// TIA Portal project "Linie_reciclare_paleti_mod" (V16)

(* hardware
DEVICE "S7-1200 station_1"  S7-1200 Station
   slot 0: "Rack_0"  S7-1200 Rack  Rack  V1.0
   slot 1: "150A19"  CPU 1214C DC/DC/Rly  6ES7 214-1HG40-0XB0  V4.4
   slot 2: "150A1101"  SM 1221 DI8 x 24VDC  6ES7 221-1BF30-0XB0  V1.0
   slot 3: "150A1102"  SM 1221 DI8 x 24VDC  6ES7 221-1BF30-0XB0  V1.0
   slot 4: "150A1103"  6ES7 221-1BH32-0XB0  V2.0
   slot 5: "150A1104"  6ES7 221-1BH32-0XB0  V2.0
   slot 6: "150A1105"  6ES7 221-1BH32-0XB0  V2.0
   slot 7: "150A1201"  SM 1222 DQ8 x relay  6ES7 222-1HF32-0XB0  V2.0
   slot 8: "150A1202"  SM 1222 DQ8 x relay  6ES7 222-1HF32-0XB0  V2.0
   slot 9: "150A1203"  SM 1222 DQ16 x relay  6ES7 222-1HH32-0XB0  V2.0
DEVICE "Master_Destacker"  GSD.Device.PN
   slot 0: "Rack"  Rack  V1.0
   slot 0: "Master_Destacker"  AL1100  AL1100
      slot 0: "AL1100"  AL1100
      slot 1: "X1"  X1
         slot 1: "Port 1"  Port 1
         slot 2: "Port 2"  Port 2
      slot 1: "4 Ports_1"  4 Ports  AL1100
         slot 0: "IO-Link Master"  IO-Link Master
   slot 1: "AL2401_IO-Link In  4 Byte + PQI"  IO-Link In  4 Byte + PQI
   slot 2: "AL2401_IO-Link In  4 Byte + PQI_1"  IO-Link In  4 Byte + PQI
   slot 3: "AL2330_IO-Link In/Out  8/ 8 Byte + PQI"  IO-Link In/Out  8/ 8 Byte + PQI
   slot 4: "IO-Link In/Out  2/ 2 Byte + PQI"  IO-Link In/Out  2/ 2 Byte + PQI
DEVICE "Master_Stacker"  GSD.Device.PN
   slot 0: "Rack"  Rack  V1.0
   slot 0: "Master_Stacker"  AL1100  AL1100
      slot 0: "AL1100"  AL1100
      slot 1: "X1"  X1
         slot 1: "Port 1"  Port 1
         slot 2: "Port 2"  Port 2
      slot 1: "4 Ports_1"  4 Ports  AL1100
         slot 0: "IO-Link Master"  IO-Link Master
   slot 1: "IO-Link In  4 Byte + PQI"  IO-Link In  4 Byte + PQI
   slot 2: "IO-Link In  4 Byte + PQI_1"  IO-Link In  4 Byte + PQI
   slot 3: "IO-Link In/Out  8/ 8 Byte + PQI"  IO-Link In/Out  8/ 8 Byte + PQI
   slot 4: "IO-Link In/Out  2/ 2 Byte + PQI"  IO-Link In/Out  2/ 2 Byte + PQI
DEVICE "HMI_1"  KTP700 Basic PN
   slot 0: "HMI_1"  KTP700 Basic PN  6AV2 123-2GB03-0AX0  16.0.0.0
   slot 1: "HMI_RT_1"  KTP700 Basic PN  6AV2 123-2GB03-0AX0  16.0.0.0
   slot 5: "HMI_1.IE_CP_1"  PROFINET Interface  16.0.0.0
      slot 1: "PROFINET Interface_1"  PROFINET Interface
         slot 1: "Port_1"  Port
DEVICE "HMI_2"  KTP700 Basic PN
   slot 0: "HMI_1"  KTP700 Basic PN  6AV2 123-2GB03-0AX0  16.0.0.0
   slot 1: "HMI_RT_2"  KTP700 Basic PN  6AV2 123-2GB03-0AX0  16.0.0.0
   slot 5: "HMI_1.IE_CP_1"  PROFINET Interface  16.0.0.0
      slot 1: "PROFINET Interface_1"  PROFINET Interface
         slot 1: "Port_1"  Port
*)

// ===== PLC "150A19"  CPU 1214C DC/DC/Rly =====

VAR_GLOBAL   // PLC tag table "Default tag table"
   "MD_IS1_SC_X1.0" AT %I70.0 : Bool;
   "MD_IS1_SC_X1.1" AT %I70.1 : Bool;
   "MD_IS1_SC_X1.2" AT %I70.2 : Bool;
   "MD_IS1_SC_X1.3" AT %I70.3 : Bool;
   "MD_IS1_SC_X1.4" AT %I70.4 : Bool;
   "MD_IS1_SC_X1.5" AT %I70.5 : Bool;
   "MD_IS1_SC_X1.6" AT %I70.6 : Bool;
   "MD_IS1_SC_X1.7" AT %I70.7 : Bool;
   "MD_IS2_SC_X1.0" AT %I75.0 : Bool;
   "MD_IS2_SC_X1.1" AT %I75.1 : Bool;
   "MD_IS2_SC_X1.2" AT %I75.2 : Bool;
   "MD_IS2_SC_X1.3" AT %I75.3 : Bool;
   "MD_IS2_SC_X1.4" AT %I75.4 : Bool;
   "MD_IS2_SC_X1.5" AT %I75.5 : Bool;
   "MD_IS2_SC_X1.6" AT %I75.6 : Bool;
   "MD_IS2_SC_X1.7" AT %I75.7 : Bool;
   "MD_OS_SC_X1.0" AT %I92.0 : Bool;
   "MD_OS_SC_X1.1" AT %I93.0 : Bool;
   "MD_OS_SC_X1.2" AT %I92.1 : Bool;
   "MD_OS_SC_X1.3" AT %I93.1 : Bool;
   "MD_OS_SC_X1.4" AT %I92.2 : Bool;
   "MD_OS_SC_X1.5" AT %I93.2 : Bool;
   "MS_IS1_SC_X1.0" AT %I80.0 : Bool;
   "MS_IS1_SC_X1.1" AT %I80.1 : Bool;
   "MS_IS1_SC_X1.2" AT %I80.2 : Bool;
   "MS_IS1_SC_X1.3" AT %I80.3 : Bool;
   "MS_IS1_SC_X1.4" AT %I80.4 : Bool;
   "MS_IS1_SC_X1.5" AT %I80.5 : Bool;
   "MS_IS1_SC_X1.6" AT %I80.6 : Bool;
   "MS_IS1_SC_X1.7" AT %I80.7 : Bool;
   "MS_IS2_SC_X1.0" AT %I85.0 : Bool;
   "MS_IS2_SC_X1.1" AT %I85.1 : Bool;
   "MS_IS2_SC_X1.2" AT %I85.2 : Bool;
   "MS_IS2_SC_X1.3" AT %I85.3 : Bool;
   "MS_IS2_SC_X1.4" AT %I85.4 : Bool;
   "MS_IS2_SC_X1.5" AT %I85.5 : Bool;
   "MS_IS2_SC_X1.6" AT %I85.6 : Bool;
   "MS_IS2_SC_X1.7" AT %I85.7 : Bool;
   "MS_OS_SC_X1.0" AT %I101.0 : Bool;
   "MS_OS_SC_X1.1" AT %I102.0 : Bool;
   "MS_OS_SC_X1.2" AT %I101.1 : Bool;
   "MS_OS_SC_X1.3" AT %I102.1 : Bool;
   "MS_OS_SC_X1.4" AT %I101.2 : Bool;
   "MS_OS_SC_X1.5" AT %I102.2 : Bool;
   "DS_AlarmMovement" AT %MW2 : Word;
   "S_AlarmMovement" AT %MW4 : Word;
   "DS_oAlarmForks" AT %M2.1 : Bool;
   "DS_oAlarmPosition" AT %M2.2 : Bool;
   "S_oAlarmUpDown" AT %M4.0 : Bool;
   "S_oAlarmForks" AT %M4.1 : Bool;
   "S_oAlarmPosition" AT %M4.2 : Bool;
   "DS_oAlarmUpDown" AT %M2.0 : Bool;
   "NOP" AT %M3.0 : Bool;
   "System_Byte" AT %MB1 : Byte;
   "FirstScan" AT %M1.0 : Bool;
   "DiagStatusUpdate" AT %M1.1 : Bool;
   "AlwaysTRUE" AT %M1.2 : Bool;
   "AlwaysFALSE" AT %M1.3 : Bool;
   "Clock_Byte" AT %MB0 : Byte;
   "Clock_10Hz" AT %M0.0 : Bool;
   "Clock_5Hz" AT %M0.1 : Bool;
   "Clock_2.5Hz" AT %M0.2 : Bool;
   "Clock_2Hz" AT %M0.3 : Bool;
   "Clock_1.25Hz" AT %M0.4 : Bool;
   "Clock_1Hz" AT %M0.5 : Bool;
   "Clock_0.625Hz" AT %M0.6 : Bool;
   "Clock_0.5Hz" AT %M0.7 : Bool;
   "M_Reset_Faults" AT %M3.1 : Bool;
   "Tag_1" AT %M3.5 : Bool;
   "Maintenance" AT %M5.0 : Bool;
   "Rez_G7_DS" AT %M6.0 : Bool;
   "Rez_G7_S" AT %M6.1 : Bool;
   "Fault_Length_DS" AT %M6.2 : Bool;
   "Fault_Length_S" AT %M6.3 : Bool;
   "Fault_Length_DS_ACK" AT %M6.4 : Bool;
   "Fault_Length_S_ACK" AT %M6.5 : Bool;
   "Length_DS_ACK" AT %M7.0 : Bool;
   "Length_S_ACK" AT %M7.2 : Bool;
   "Length_DS_HMI_1" AT %M14.0 : Bool;
   "Length_DS_HMI_2" AT %M14.1 : Bool;
   "Length_DS_HMI_3" AT %M14.2 : Bool;
   "Length_S_HMI_1" AT %M14.3 : Bool;
   "Length_S_HMI_2" AT %M14.4 : Bool;
   "Length_S_HMI_3" AT %M14.5 : Bool;
   "Manual_Reset Destacker 110KF1 Safety Relay" AT %M8.0 : Bool;
   "Manual_Reset Destacker 111KF1 Safety Barrier Relay" AT %M8.1 : Bool;
   "Manual_Reset Zone 2 112KF1 Safety Relay" AT %M8.2 : Bool;
   "Manual_Reset Stacker 113KF1 Safety Relay" AT %M8.3 : Bool;
   "Manual_Reset Stacker 114KF1 Safety Barrier Relay 1" AT %M8.4 : Bool;
   "Manual_Reset Stacker 115KF1 Safety Barrier Relay 2" AT %M8.5 : Bool;
   "Manual_Cuplare contactor VFD Conveior 1 alimentare destacker" AT %M8.6 : Bool;
   "Manual_ON/OFF1 VFD Conveior 1 alimentare destacker" AT %M8.7 : Bool;
   "Manual_Fault Aknowledge VFD Conveior 1 alimentare destacker" AT %M9.0 : Bool;
   "Manual_Cuplare contactor VFD Conveior 2 iesire destacker" AT %M9.1 : Bool;
   "Manual_ON/OFF1 VFD Conveior 2 iesire destacker" AT %M9.2 : Bool;
   "Manual_Fault Aknowledge VFD Conveior 2 iesire destacker" AT %M9.3 : Bool;
   "Manual_Start Conveior 1 preluare paleti OK" AT %M9.4 : Bool;
   "Manual_Softstarter aer 1.1 Conveior 1 preluare paleti OK" AT %M9.5 : Bool;
   "Manual_Softstarter aer 1.2 Conveior 1 preluare paleti OK" AT %M9.6 : Bool;
   "Manual_Start Conveior 2 transfer palet 1" AT %M9.7 : Bool;
   "Manual_Cuplare contactor VFD Conveior 3 transfer palet 2" AT %M10.0 : Bool;
   "Manual_ON/OFF1 VFD Conveior 3 transfer palet 2" AT %M10.1 : Bool;
   "Manual_Fault Aknowledge VFD Conveior 3 transfer palet 2" AT %M10.2 : Bool;
   "Manual_Cuplare contactor VFD Conveior 4 descarcare stacker" AT %M10.3 : Bool;
   "Manual_ON/OFF1 VFD Conveior 4 descarcare stacker" AT %M10.4 : Bool;
   "Manual_Fault Aknowledge VFD Conveior 4 descarcare stacker" AT %M10.5 : Bool;
   "Manual_DS_Comanda cilindru vertical sus" AT %M10.6 : Bool;
   "Manual_DS_Comanda cilindru vertical jos" AT %M10.7 : Bool;
   "Manual_DS_Comanda furca retrasa" AT %M11.0 : Bool;
   "Manual_Comanda 1 softstarter aer destacker" AT %M11.1 : Bool;
   "Manual_Comanda 2 softstarter aer destacker" AT %M11.2 : Bool;
   "Manual_Feed palet (LED temp)" AT %M11.3 : Bool;
   "Manual_S_Comanda cilindru vertical sus" AT %M11.4 : Bool;
   "Manual_S_Comanda cilindru vertical jos" AT %M11.5 : Bool;
   "Manual_S_Comanda furca extinsa" AT %M11.6 : Bool;
   "Manual_S_Comanda furca retrasa" AT %M11.7 : Bool;
   "Manual_Comanda 1 softstarter aer stacker" AT %M12.0 : Bool;
   "Manual_Comanda 2 softstarter aer stacker" AT %M12.1 : Bool;
   "Manual_Comanda intrare cilindru centrare" AT %M12.2 : Bool;
   "Manual_Comanda iesire cilindru centrare" AT %M12.3 : Bool;
   "Manual_DS_Comanda furca extinsa" AT %M12.4 : Bool;
   "No_Safe_DS" AT %M13.0 : Bool;
   "Energie_SN" AT %M13.1 : Bool;
   "Manual_DS" AT %M13.2 : Bool;
   "Automat_DS" AT %M13.3 : Bool;
   "Wait_Start_Cycle_DS" AT %M13.4 : Bool;
   "Cycle_Run_DS" AT %M13.5 : Bool;
   "Init_DS" AT %M13.6 : Bool;
   "Init_Done_DS" AT %M13.7 : Bool;
   "Safe_SN" AT %M14.6 : Bool;
   "No_Safe_S" AT %M14.7 : Bool;
   "Energie_S" AT %M15.0 : Bool;
   "Manual_S" AT %M15.1 : Bool;
   "Automat_S" AT %M15.2 : Bool;
   "Wait_Start_Cycle_S" AT %M15.3 : Bool;
   "Cycle_Run_S" AT %M15.4 : Bool;
   "Init_S" AT %M15.5 : Bool;
   "Init_Done_S" AT %M15.6 : Bool;
   "Safe_S" AT %M15.7 : Bool;
   "Alarm_Stop_DS" AT %M16.0 : Bool;
   "bStop_DS" AT %M16.1 : Bool;
   "Alarm_Stop_S" AT %M16.2 : Bool;
   "bStop_S" AT %M16.3 : Bool;
   "Centrat" AT %M16.4 : Bool;
   "td" AT %M6.6 : Bool;
   "NoTranzit" AT %M7.3 : Bool;
   "NoCylAdv" AT %M6.7 : Bool;
   "NoProd" AT %M7.1 : Bool;
   "ForceIniCylRet" AT %M17.0 : Bool;
   "RstAlm" AT %M7.4 : Bool;
   "ForceIniTranzit" AT %M7.5 : Bool;
   "ForceIniProdus" AT %M7.6 : Bool;
   "bStart_DS" AT %M12.5 : Bool;
   "bStart_S" AT %M7.7 : Bool;
   "bStepper_S" AT %M12.6 : Bool;
   "bStepper_DS" AT %M12.7 : Bool;
   "Safe_Z2_A" AT %M16.6 : Bool;
   "Energie_Z2_A" AT %M16.5 : Bool;
   "Home_S" AT %M16.7 : Bool;
   "Extins_Recul_Mem" AT %M17.1 : Bool;
   "CPO_Sim" AT %M97.0 : Bool;
   "ForceTim" AT %M17.2 : Bool;
   "b0" AT %M17.3 : Bool;
   "RstAlmF" AT %M17.4 : Bool;
   "TrigChart" AT %M17.5 : Bool;
   "SCentrorMem" AT %M17.6 : Bool;
   "SCentrorMemT" AT %M17.7 : Bool;
   "Cycle_Run_Palet" AT %M18.0 : Bool;
   "DeliveryNew" AT %M18.1 : Bool;
   "req_evac" AT %M18.2 : Bool;
   "fr" AT %M18.3 : Bool;
   "ChgLowSpd" AT %M18.4 : Bool;
   "ChgLowSpd_pre" AT %M18.5 : Bool;
   "S_actMut" AT %M18.6 : Bool;
   "StopCmdDn1" AT %M19.0 : Bool;
   "StopCmdDn2" AT %M19.2 : Bool;
   "SkipSenzor" AT %M18.7 : Bool;
   "Home_SN" AT %M19.3 : Bool;
   "Fault_Length_SN" AT %M19.1 : Bool;
   "SNCentrorMem" AT %M19.4 : Bool;
   "SNCentrorMemT" AT %M19.5 : Bool;
   "Automat_SN" AT %M19.6 : Bool;
   "Init_SN" AT %M19.7 : Bool;
   "bStepper_SN" AT %M20.0 : Bool;
   "bStop_SN" AT %M20.1 : Bool;
   "bStart_SN" AT %M20.2 : Bool;
   "SN_actMut" AT %M20.3 : Bool;
   "SNChgLowSpd" AT %M20.4 : Bool;
   "SNChgLowSpd_pre" AT %M20.5 : Bool;
   "SN_fr" AT %M20.6 : Bool;
   "SN_req_evac" AT %M20.7 : Bool;
   "SN_Cycle_Run_Palet" AT %M21.0 : Bool;
   "SN_NoCylAdv" AT %M21.1 : Bool;
   "SN_NoProd" AT %M21.2 : Bool;
   "SN_NoTranzit" AT %M21.3 : Bool;
   "SN_DeliveryNew" AT %M21.4 : Bool;
END_VAR

VAR_GLOBAL   // PLC tag table "150A19"
   "110KF1" AT %I0.0 : Bool;   // E-Stop Line B 110KF1 Safety Relay
   "111KF1" AT %I0.1 : Bool;   // Stacker Nou 111KF1 Safety Barrier Relay Mutting
   "112KF1" AT %I0.2 : Bool;   // E-Stop Line A 112KF1 Safety Relay
   "113KF1" AT %I0.3 : Bool;   // Stacker 113KF1 Safety Relay
   "114KF1" AT %I0.4 : Bool;   // Stacker 114KF1 Safety Barrier Relay 1
   "115KF1" AT %I0.5 : Bool;   // Stacker 115KF1 Safety Barrier Relay Mutting
   "110S1" AT %I0.6 : Bool;   // Emergency Stop Stacker Nou
   "112S1" AT %I0.7 : Bool;   // Emergency Stop Zone 2_A
   "113S1" AT %I1.0 : Bool;   // Emergency Stop Stacker
   "155S1" AT %I1.1 : Bool;   // Reset safety General
   "151S1" AT %I2.0 : Bool;   // Prezenta aer
   "105F2" AT %I2.1 : Bool;   // Protectie cuplata Iluminat
   "120Q1" AT %I2.2 : Bool;   // Protectie cuplata Conveior 1 alimentare stacker nou
   "121K1" AT %I2.3 : Bool;   // Contactor cuplat Conveior 1 alimentare stacker nou
   "120K1" AT %I2.4 : Bool;   // Frana decuplata Conveior 1 alimentare stacker nou
   "120U1_PowerOK" AT %I2.5 : Bool;   // Functionare Conveior 1 alimentare stacker nou
   "120U1_Fault" AT %I2.6 : Bool;   // Avarie Conveior 1 alimentare stacker nou
   "122Q1" AT %I2.7 : Bool;   // Protectie cuplata Conveior 2 iesire stacker nou
   "123K1" AT %I3.0 : Bool;   // Contactor cuplat Conveior 2 iesire stacker nou
   "122K1" AT %I3.1 : Bool;   // Frana decuplata Conveior 2 iesire stacker nou
   "122U1_PowerOK" AT %I3.2 : Bool;   // Functionare Conveior 2 iesire stacker nou
   "122U1_Fault" AT %I3.3 : Bool;   // Avarie Conveior 2 iesire stacker nou
   "124Q1" AT %I3.4 : Bool;   // Protectie cuplata Conveior 1 preluare paleti OK Zona A
   "124K1" AT %I3.5 : Bool;   // Functionare Conveior 1 preluare paleti OK Zona A
   "125Q1" AT %I3.6 : Bool;   // Protectie cuplata Conveior 2 transfer palet 1 Zona A
   "125K1" AT %I3.7 : Bool;   // Functionare Conveior 2 transfer palet 1 Zona A
   "126Q1" AT %I4.0 : Bool;   // Protectie cuplata Conveior 3 transfer palet 2
   "127K1" AT %I4.1 : Bool;   // Contactor cuplat Conveior 3 transfer palet 2
   "126K1" AT %I4.2 : Bool;   // Frana decuplata Conveior 3 transfer palet 2
   "126U1_PowerOK" AT %I4.3 : Bool;   // Functionare Conveior 3 transfer palet 2
   "126U1_Fault" AT %I4.4 : Bool;   // Avarie Conveior 3 transfer palet 2
   "128Q1" AT %I4.5 : Bool;   // Protectie cuplata Conveior 4 descarcare stacker
   "129K1" AT %I4.6 : Bool;   // Contactor cuplat Conveior 4 descarcare stacker
   "128K1" AT %I4.7 : Bool;   // Frana decuplata Conveior 4 descarcare stacker
   "128U1_PowerOK" AT %I5.0 : Bool;   // Functionare Conveior 4 stacker
   "128U1_Fault" AT %I5.1 : Bool;   // Avarie Conveior 4 stacker
   "102F1" AT %I5.2 : Bool;   // Protectie cuplata Masina demontare paleti stanga
   "103F1" AT %I5.3 : Bool;   // Protectie cuplata Masina demontare paleti dreapta
   "104F1" AT %I5.4 : Bool;   // Protectie cuplata Circular masa fixa
   "105F1" AT %I5.5 : Bool;   // Protectie cuplata Post reparatie stanga+dreapta
   "106F1" AT %I5.6 : Bool;   // Protectie cuplata Post reparatii minore
   "107F1" AT %I5.7 : Bool;   // Protectie cuplata TELE
   "149F1" AT %I7.0 : Bool;   // Protectie cuplata HMI
   "141VFA1_SQ1" AT %I7.1 : Bool;   // Senzor 1 proximitate softstarter aer zona 2 A
   "141VFA1_SQ2" AT %I7.2 : Bool;   // Senzor 2 proximitate softstarter aer zona 2 A
   "124Q2" AT %I7.3 : Bool;   // Protectie cuplata Conveior 1 preluare paleti OK Zona B
   "Puls_Consum" AT %I7.4 : Bool;
   "124K2" AT %I7.5 : Bool;   // Functionare Conveior 1 preluare paleti OK Zona B
   "125Q2" AT %I7.6 : Bool;   // Protectie cuplata Conveior 2 transfer palet 1 Zona B
   "125K2" AT %I7.7 : Bool;   // Functionare Conveior 2 transfer palet 1 Zona B
   "153K1" AT %Q0.0 : Bool;   // Reset stacker nou 110KF1 Safety Relay
   "153K2" AT %Q0.1 : Bool;   // Reset stacker nou 111KF1 Safety Barrier Relay
   "153K3" AT %Q0.2 : Bool;   // Reset Zone 2 112KF1 Safety Relay
   "153K4" AT %Q0.3 : Bool;   // Reset Stacker 113KF1 Safety Relay
   "153K5" AT %Q0.4 : Bool;   // Reset Stacker 114KF1 Safety Barrier Relay 1
   "153K6" AT %Q0.5 : Bool;   // Reset Stacker 115KF1 Safety Barrier Relay 2
   "BD_R" AT %Q0.6 : Bool;   // S_Baliza dulap rosu
   "BD_G" AT %Q0.7 : Bool;   // S_Baliza dulap verde
   "SN_Comanda cilindru centrare" AT %Q9.6 : Bool;   // SN_Comanda cilindru centrare
   "SN_Comanda ELIBERARE cilindru centrare" AT %Q9.7 : Bool;   // SN_Comanda ELIBERARE cilindru centrare
   "CSN3_PowerOK" AT %Q7.3 : Bool;   // SN_Cuplare contactor VFD Conveior 1 alimentare
   "CSN3_Start" AT %Q7.4 : Bool;   // SN_ON/OFF1 VFD Conveior 1 alimentare
   "CSN4_PowerOK" AT %Q7.5 : Bool;   // SN_Cuplare contactor VFD Conveior 2 iesire
   "CSN4_Start" AT %Q7.6 : Bool;   // SN_ON/OFF1 VFD Conveior 2 iesire
   "CS1_Start" AT %Q8.0 : Bool;   // S_Start Conveior 1 preluare paleti OK
   "Softstarter aer 1.1 Conveior 1 preluare paleti OK" AT %Q8.1 : Bool;   // Softstarter aer 1.1 Conveior 1 preluare paleti OK
   "Softstarter aer 1.2 Conveior 1 preluare paleti OK" AT %Q8.2 : Bool;   // Softstarter aer 1.2 Conveior 1 preluare paleti OK
   "CS2_Start" AT %Q7.0 : Bool;   // S_Start Conveior 2 transfer palet 1
   "CS3_PowerOK" AT %Q8.3 : Bool;   // Cuplare contactor VFD Conveior 3 transfer palet 2
   "CS3_Start" AT %Q8.4 : Bool;   // ON/OFF1 VFD Conveior 3 transfer palet 2
   "CS4_PowerOK" AT %Q8.5 : Bool;   // Cuplare contactor VFD Conveior 4 descarcare stacker
   "CS4_Start" AT %Q8.6 : Bool;   // ON/OFF1 VFD Conveior 4 descarcare stacker
   "CSN2_Start" AT %Q9.0 : Bool;   // SN_Start Conveior 2 transfer palet 1
   "CSN1_Start" AT %Q9.3 : Bool;   // SN_Start Conveior 2 transfer palet 1
   "Comanda 1 softstarter aer Zona B" AT %Q9.4 : Bool;   // Comanda 1 softstarter aer Zona B
   "Comanda 2 softstarter aer Zona B" AT %Q9.5 : Bool;   // Comanda 2 softstarter aer Zona B
   "S_Comanda cilindru centrare" AT %Q7.1 : Bool;   // S_Comanda cilindru centrare
   "S_Comanda ELIBERARE cilindru centrare" AT %Q7.2 : Bool;   // S_Comanda ELIBERARE cilindru centrare
   "CS3_SlowSpeed" AT %Q8.7 : Bool;   // Slow speed
   "CSN3_SlowSpeed" AT %Q7.7 : Bool;   // Slow speed
   "StopInUp1" AT %I6.0 : Bool;   // StopInUp1
   "StopInDn1" AT %I6.1 : Bool;   // StopInDn1
   "StopInUp2" AT %I6.2 : Bool;   // StopInUp2
   "StopInDn2" AT %I6.3 : Bool;   // StopInDn2
   "S_ActMutting" AT %Q1.0 : Bool;   // Activare Muting Stacker
   "SN_ActMutting" AT %Q1.1 : Bool;   // Activare Muting Stacker Nou
   "CSN3_FaultAck" AT %Q10.0 : Bool;   // SN_Fault Aknowledge VFD Conveior 1 alimentare
   "CSN4_FaultAck" AT %Q10.1 : Bool;   // SN_Fault Aknowledge VFD Conveior 2 iesire
   "CS3_FaultAck" AT %Q10.2 : Bool;   // Fault Aknowledge VFD Conveior 3 transfer palet 2
   "StopCmdUp2" AT %Q10.4 : Bool;
   "StopCmdUp1" AT %Q10.5 : Bool;
   "CS4_FaultAck" AT %Q10.3 : Bool;   // Fault Aknowledge VFD Conveior 4 descarcare stacker
   "SN_Baliza dulap rosu" AT %M21.5 : Bool;
   "Sn_Baliza dulap verde" AT %M21.6 : Bool;
   "114S1" AT %I1.2 : Bool;   // Emergency Stop Zone 2_B
   "Safe_Z2_B" AT %M21.7 : Bool;
   "100KF1" AT %I1.3 : Bool;   // Safety Relay Main Door
   "142VFA1_SQ2" AT %I6.5 : Bool;   // Senzor 2 proximitate softstarter aer zona 2 B
   "142VFA1_SQ1" AT %I6.4 : Bool;   // Senzor 1 proximitate softstarter aer zona 2 B
   "Energie_Z2_B" AT %M22.0 : Bool;
   "ngr" AT %M22.1 : Bool;
END_VAR

VAR_GLOBAL   // PLC tag table "160A19"
   "CSN1_SQ1" AT %I68.0 : Bool;   // SN_Prezenta palet
   "CSN1_SQ3" AT %I68.1 : Bool;   // SN_Prezenta palet_capat_conveyor
   "CSN2_SQ1" AT %I68.2 : Bool;   // SN_Masurare lungime
   "CSN3_SQ2" AT %I68.3 : Bool;   // SN_Lungime 2
   "CSN4_SQ1" AT %I68.4 : Bool;   // SN_Prezenta stiva
   "CPN2_SQ2" AT %I68.5 : Bool;   // SN_Centror retras
   "1XXS2" AT %I68.6 : Bool;   // SN_Reset safety Stacker_New
   "SN_Prezenta palet_centror" AT %I69.1 : Bool;   // SN_Prezenta palet_centror
   "CSN3_SQ1" AT %I69.2 : Bool;   // SN_Lungime 1
   "CSN3_SQ3" AT %I69.3 : Bool;   // SN_Lungime 3
   "SN_Switch_Iesire" AT %I69.4 : Bool;   // SN_Switch_Iesire
   "CPN2_SQ3" AT %I69.5 : Bool;   // SN_Centror extins
   "SN_Prez_conveyor_volum" AT %I69.6 : Bool;   // SN_Prez_conveyor_volum
   "SN_Senzor stacking" AT %I73.1 : Bool;   // SN_Senzor stacking
   "SN_Cilindru vertical sus" AT %I73.2 : Bool;   // SN_Cilindru vertical sus
   "SN_Cilindru vertical mijloc" AT %I73.3 : Bool;   // SN_Cilindru vertical mijloc
   "SN_Detectie palet" AT %I73.4 : Bool;   // SN_Detectie palet
   "SN_Cilindru vertical jos" AT %I73.5 : Bool;   // SN_Cilindru vertical jos
   "SN_Cilindru retras" AT %I74.1 : Bool;   // SN_Cilindru retras
   "SN_Cilindru extins" AT %I74.6 : Bool;   // SN_Cilindru extins
   "SN_Furca_liber1" AT %I73.0 : Bool;   // SN_Furca_liber1
   "SN_Furca_liber2" AT %I74.0 : Bool;   // SN_Furca_liber2
   "SN_Reset safety Stacker_2" AT %I73.6 : Bool;   // SN_Reset safety Stacker_2
   "140VFA1_SQ1" AT %I73.7 : Bool;   // Senzor 1 proximitate softstarter aer stacker nou
   "140VFA1_SQ2" AT %I74.7 : Bool;   // Senzor 2 proximitate softstarter aer stacker nou
   "BSN_R" AT %Q3.0 : Bool;   // BDS_R
   "BSN_G" AT %Q3.1 : Bool;   // BDS_G
   "BSN_Y" AT %Q3.3 : Bool;   // BDS_Y
   "SN_Comanda cilindru vertical sus" AT %Q64.0 : Bool;   // SN_Comanda cilindru vertical sus
   "Comanda 1 softstarter aer stacker_new" AT %Q64.1 : Bool;   // Comanda 1 softstarter aer stacker_new
   "SN_Comanda furca retrasa" AT %Q65.0 : Bool;   // SN_Comanda furca retrasa
   "SN_Comanda cilindru vertical jos" AT %Q66.0 : Bool;   // SN_Comanda cilindru vertical jos
   "Comanda 2 softstarter aer stacker_new" AT %Q66.1 : Bool;   // Comanda 2 softstarter aer stacker_new
   "SN_Comanda furca extinsa" AT %Q67.0 : Bool;   // SN_Comanda furca extinsa
   "Door_Left Open" AT %I69.0 : Bool;
END_VAR

VAR_GLOBAL   // PLC tag table "180A19"
   "CS1_SQ1" AT %I78.0 : Bool;   // S_Prezenta palet
   "CS1_SQ3" AT %I78.1 : Bool;   // S_Prezenta palet_capat_conveyor
   "CS2_SQ1" AT %I78.2 : Bool;   // S_Masurare lungime
   "CS3_SQ2" AT %I78.3 : Bool;   // S_Lungime 2
   "CS4_SQ1" AT %I78.4 : Bool;   // S_Prezenta_stiva
   "CP2_SQ2" AT %I78.5 : Bool;   // S_Centror retras
   "110S2" AT %I78.6 : Bool;   // S_Reset safety Stacker
   "CS3_SQ1" AT %I79.2 : Bool;   // S_Lungime 1
   "CS3_SQ3" AT %I79.3 : Bool;   // S_Lungime 3
   "CP2_SQ3" AT %I79.5 : Bool;   // S_Centror extins
   "S_Prezenta palet_centror" AT %I79.1 : Bool;   // S_Prezenta palet_centror
   "S_Switch_iesire" AT %I79.4 : Bool;   // S_Switch_iesire
   "S_Prez_conveyor_volum" AT %I78.7 : Bool;   // S_Prez_conveyor_volum
   "S_Furca_liber1" AT %I83.0 : Bool;   // S_Furca_liber1
   "S_Senzor stacking" AT %I83.1 : Bool;   // S_Senzor stacking
   "S_Cilindru vertical sus" AT %I83.2 : Bool;   // S_Cilindru vertical sus
   "S_Cilindru vertical mijloc" AT %I83.3 : Bool;   // S_Cilindru vertical mijloc
   "S_Detectie palet" AT %I83.4 : Bool;   // S_Detectie palet
   "S_Cilindru vertical jos" AT %I83.5 : Bool;   // S_Cilindru vertical jos
   "S_Reset safety Stacker_2" AT %I83.6 : Bool;   // S_Reset safety Stacker_2
   "143VFA1_SQ1" AT %I83.7 : Bool;   // S_Senzor 1 proximitate softstarter aer stacker
   "S_Furca_liber2" AT %I84.0 : Bool;   // S_Furca_liber2
   "S_Cilindru retras" AT %I84.1 : Bool;   // S_Cilindru retras
   "S_Cilindru extins" AT %I84.6 : Bool;   // S_Cilindru extins
   "143VFA1_SQ2" AT %I84.7 : Bool;   // S_Senzor 2 proximitate softstarter aer stacker
   "BS_R" AT %Q13.0 : Bool;   // S_BS_R
   "BS_G" AT %Q13.1 : Bool;   // S_BS_G
   "BS_Y" AT %Q13.3 : Bool;   // S_BS_Y
   "S_Comanda cilindru vertical sus" AT %Q72.0 : Bool;   // S_Comanda cilindru vertical sus
   "Comanda 1 softstarter aer stacker" AT %Q72.1 : Bool;   // Comanda 1 softstarter aer stacker
   "S_Comanda furca retrasa" AT %Q73.0 : Bool;   // S_Comanda furca retrasa
   "S_Comanda cilindru vertical jos" AT %Q74.0 : Bool;   // S_Comanda cilindru vertical jos
   "Comanda 2 softstarter aer stacker" AT %Q74.1 : Bool;   // Comanda 2 softstarter aer stacker
   "S_Comanda furca extinsa" AT %Q75.0 : Bool;   // S_Comanda furca extinsa
   "Door_Front Open" AT %I79.0 : Bool;
END_VAR

TYPE "OP_Int"
VERSION : 0.1
   STRUCT
      O_ComActive : Bool;
      O_Fault : Bool;
      I_DataStorage : Bool;
      I_BlockParam : Bool;
      IO_ReadReq : Bool;
      IO_WriteReq : Bool;
      IO_Ackn : Bool;
      IO_EventRead : Bool;
      IO_ParamConfigFaultRead : Bool;
   END_STRUCT;
END_TYPE

TYPE "udt_station"
VERSION : 0.1
   STRUCT
      mpp : Bool;
      ip : Bool;
      alm_apar : Bool;
      alar_disapear : Bool;
      alm_tmt : Bool;
      alm_release : Bool;
      AuthAdmit : Bool;
      almt : Bool;
      WrkDn : Bool;
      "step" : USInt;
      stepv : USInt;
      test : USInt;
      alm_tim : Array[1..6] of IEC_TIMER;
   END_STRUCT;
END_TYPE

TYPE "PQI_IF"
VERSION : 0.1
   STRUCT
      O_DI4 : Bool;
      O_DI2 : Bool;
      O_DA : Bool;
      O_DE : Bool;
      O_PQ : Bool;
   END_STRUCT;
END_TYPE

TYPE "Bits_Destacker"
VERSION : 0.1
   STRUCT
      Input : Struct
         iEnable : Bool;
         iReset : Bool;
         iAutomatic : Bool;
         iManual : Bool;
         iManualUp : Bool;
         iManualDown : Bool;
         iManualOpenForks : Bool;
         iManualCloseForks : Bool;
         Vertical_sus : Bool;
         Vertical_mijloc : Bool;
         iB10 : Bool;
         Vertical_jos : Bool;
         Furca_extins : Bool;
         Furca_retras : Bool;
         Detectie_palet : Bool;
         Senzor_stiva : Bool;
      END_STRUCT;
      Output : Struct
         Cmd_sus : Bool;
         Cmd_jos : Bool;
         Cmd_extindere : Bool;
         Cmd_retragere : Bool;
         oAlarmUpDown : Bool;
         oAlarmForks : Bool;
         oAlarmPosition : Bool;
         oAlarmEmpty : Bool;
         oAlarmAlmostEmpty : Bool;
      END_STRUCT;
   END_STRUCT;
END_TYPE

TYPE "IF_AL2401"
VERSION : 0.1
   STRUCT
      StandardStructure : Struct
         Header : Struct
            NumberParameter : Int := 15;
            AdressParamDownLoad : Int := 20;
            AdressDeviceIndent : Int := 44;
            AdressApplicSpez : Int := 700;
            AdressDeviceParam : Int := 946;
            AdressKommando : Int := 1026;
            NumberCommandos : Int := 5;
            Spare01 : Int;
            Spare02 : Int;
            Spare03 : Int;
         END_STRUCT;
         Paramdownload : Struct
            ParamDownLoadStart : Struct
               BlockStat : DWord;
               IOLStat : DWord;
            END_STRUCT;
            ParamDownLoadEnd : Struct
               BlockStat : DWord;
               IOLStat : DWord;
            END_STRUCT;
            ParamDownLoadStore : Struct
               BlockStat : DWord;
               IOLStat : DWord;
            END_STRUCT;
         END_STRUCT;
         DeviceIndentification : Struct
            V_VendorName : Struct
               Text : String[64];
               Index : Int := 16;
               Subindex : Int := 0;
               Length : Int := 19;
               BlockStat : DWord;
               IOLStat : DWord;
               RelRead : Bool := TRUE;
               RelWrite : Bool := FALSE;
            END_STRUCT;
            V_VendorText : Struct
               Text : String[64];
               Index : Int := 17;
               Subindex : Int := 0;
               Length : Int := 11;
               BlockStat : DWord;
               IOLStat : DWord;
               RelRead : Bool := TRUE;
               RelWrite : Bool := FALSE;
            END_STRUCT;
            V_ProductName : Struct
               Text : String[64];
               Index : Int := 18;
               Subindex : Int := 0;
               Length : Int := 6;
               BlockStat : DWord;
               IOLStat : DWord;
               RelRead : Bool := TRUE;
               RelWrite : Bool := FALSE;
            END_STRUCT;
            V_ProductID : Struct
               Text : String[64];
               Index : Int := 19;
               Subindex : Int := 0;
               Length : Int := 6;
               BlockStat : DWord;
               IOLStat : DWord;
               RelRead : Bool := TRUE;
               RelWrite : Bool := FALSE;
            END_STRUCT;
            V_ProductText : Struct
               Text : String[64];
               Index : Int := 20;
               Subindex : Int := 0;
               Length : Int := 28;
               BlockStat : DWord;
               IOLStat : DWord;
               RelRead : Bool := TRUE;
               RelWrite : Bool := FALSE;
            END_STRUCT;
            V_SerialNumber : Struct
               Text : String[64];
               Index : Int := 21;
               Subindex : Int := 0;
               Length : Int := 12;
               BlockStat : DWord;
               IOLStat : DWord;
               RelRead : Bool := TRUE;
               RelWrite : Bool := FALSE;
            END_STRUCT;
            V_HardwareRevision : Struct
               Text : String[64];
               Index : Int := 22;
               Subindex : Int := 0;
               Length : Int := 2;
               BlockStat : DWord;
               IOLStat : DWord;
               RelRead : Bool := TRUE;
               RelWrite : Bool := FALSE;
            END_STRUCT;
            V_FirmwareRevision : Struct
               Text : String[64];
               Index : Int := 23;
               Subindex : Int := 0;
               Length : Int := 5;
               BlockStat : DWord;
               IOLStat : DWord;
               RelRead : Bool := TRUE;
               RelWrite : Bool := FALSE;
            END_STRUCT;
         END_STRUCT;
         ApplicationSpecificTag : Struct
            V_ApplicationSpecificTag : Struct
               Text : String[64];
               Index : Int := 24;
               Subindex : Int := 0;
               Length : Int := 32;
               BlockStat : DWord;
               IOLStat : DWord;
               RelRead : Bool := TRUE;
               RelWrite : Bool := TRUE;
            END_STRUCT;
            V_FunctionTag : Struct
               Text : String[64];
               Index : Int := 25;
               Subindex : Int := 0;
               Length : Int := 0;
               BlockStat : DWord;
               IOLStat : DWord;
               RelRead : Bool := FALSE;
               RelWrite : Bool := FALSE;
            END_STRUCT;
            V_LocationTag : Struct
               Text : String[64];
               Index : Int := 26;
               Subindex : Int := 0;
               Length : Int := 0;
               BlockStat : DWord;
               IOLStat : DWord;
               RelRead : Bool := FALSE;
               RelWrite : Bool := FALSE;
            END_STRUCT;
         END_STRUCT;
         DeviceParameters : Struct
            Parameter_01 : Struct
               V_DeviceAccessLocks : Int := 0;
               Byte02 : Byte := BYTE#16#00;
               Byte03 : Byte := BYTE#16#00;
               Index : Int := 12;
               Subindex : Int := 0;
               Length : Int := 2;
               BlockStat : DWord;
               IOLStat : DWord;
               RelRead : Bool := TRUE;
               RelWrite : Bool := TRUE;
            END_STRUCT;
            Parameter_02 : Struct
               V_DeviceStatus : Byte := BYTE#16#00;
               Byte01 : Byte := BYTE#16#00;
               Byte02 : Byte := BYTE#16#00;
               Byte03 : Byte := BYTE#16#00;
               Index : Int := 36;
               Subindex : Int := 0;
               Length : Int := 1;
               BlockStat : DWord;
               IOLStat : DWord;
               RelRead : Bool := TRUE;
               RelWrite : Bool := FALSE;
            END_STRUCT;
            Parameter_03 : Struct
               V_ShortCircuits : Int := 0;
               Byte02 : Byte := BYTE#16#00;
               Byte03 : Byte := BYTE#16#00;
               Index : Int := 687;
               Subindex : Int := 0;
               Length : Int := 2;
               BlockStat : DWord;
               IOLStat : DWord;
               RelRead : Bool := TRUE;
               RelWrite : Bool := FALSE;
            END_STRUCT;
            Parameter_04 : Struct
               V_EquipmentSpecificID : Byte := BYTE#16#00;
               Byte01 : Byte := BYTE#16#00;
               Byte02 : Byte := BYTE#16#00;
               Byte03 : Byte := BYTE#16#00;
               Index : Int := 688;
               Subindex : Int := 0;
               Length : Int := 1;
               BlockStat : DWord;
               IOLStat : DWord;
               RelRead : Bool := TRUE;
               RelWrite : Bool := TRUE;
            END_STRUCT;
         END_STRUCT;
         Commando : Struct
            Commando_00 : Struct
               Value : Byte := BYTE#16#82;
               Index : Int := 2;
               Subindex : Int := 0;
               Length : Int := 1;
               BlockStat : DWord;
               IOLStat : DWord;
            END_STRUCT;
            Commando_01 : Struct
               Value : Byte := BYTE#16#F0;
               Index : Int := 2;
               Subindex : Int := 0;
               Length : Int := 1;
               BlockStat : DWord;
               IOLStat : DWord;
            END_STRUCT;
            Commando_02 : Struct
               Value : Byte := BYTE#16#F1;
               Index : Int := 2;
               Subindex : Int := 0;
               Length : Int := 1;
               BlockStat : DWord;
               IOLStat : DWord;
            END_STRUCT;
            Commando_03 : Struct
               Value : Byte := BYTE#16#F2;
               Index : Int := 2;
               Subindex : Int := 0;
               Length : Int := 1;
               BlockStat : DWord;
               IOLStat : DWord;
            END_STRUCT;
            Commando_04 : Struct
               Value : Byte := BYTE#16#F3;
               Index : Int := 2;
               Subindex : Int := 0;
               Length : Int := 1;
               BlockStat : DWord;
               IOLStat : DWord;
            END_STRUCT;
         END_STRUCT;
      END_STRUCT;
   END_STRUCT;
END_TYPE

TYPE "IF_AL2230_AL2330"
VERSION : 0.1
   STRUCT
      StandardStructure : Struct
         Header : Struct
            NumberParameter : Int := 48;
            AdressParamDownLoad : Int := 20;
            AdressDeviceIndent : Int := 44;
            AdressApplicSpez : Int := 700;
            AdressDeviceParam : Int := 946;
            AdressKommando : Int := 1686;
            NumberCommandos : Int := 7;
            Spare01 : Int;
            Spare02 : Int;
            Spare03 : Int;
         END_STRUCT;
         Paramdownload : Struct
            ParamDownLoadStart : Struct
               BlockStat : DWord;
               IOLStat : DWord;
            END_STRUCT;
            ParamDownLoadEnd : Struct
               BlockStat : DWord;
               IOLStat : DWord;
            END_STRUCT;
            ParamDownLoadStore : Struct
               BlockStat : DWord;
               IOLStat : DWord;
            END_STRUCT;
         END_STRUCT;
         DeviceIndentification : Struct
            V_VendorName : Struct
               Text : String[64];
               Index : Int := 16;
               Subindex : Int := 0;
               Length : Int := 19;
               BlockStat : DWord;
               IOLStat : DWord;
               RelRead : Bool := TRUE;
               RelWrite : Bool := FALSE;
            END_STRUCT;
            V_VendorText : Struct
               Text : String[64];
               Index : Int := 17;
               Subindex : Int := 0;
               Length : Int := 11;
               BlockStat : DWord;
               IOLStat : DWord;
               RelRead : Bool := TRUE;
               RelWrite : Bool := FALSE;
            END_STRUCT;
            V_ProductName : Struct
               Text : String[64];
               Index : Int := 18;
               Subindex : Int := 0;
               Length : Int := 6;
               BlockStat : DWord;
               IOLStat : DWord;
               RelRead : Bool := TRUE;
               RelWrite : Bool := FALSE;
            END_STRUCT;
            V_ProductID : Struct
               Text : String[64];
               Index : Int := 19;
               Subindex : Int := 0;
               Length : Int := 6;
               BlockStat : DWord;
               IOLStat : DWord;
               RelRead : Bool := TRUE;
               RelWrite : Bool := FALSE;
            END_STRUCT;
            V_ProductText : Struct
               Text : String[64];
               Index : Int := 20;
               Subindex : Int := 0;
               Length : Int := 14;
               BlockStat : DWord;
               IOLStat : DWord;
               RelRead : Bool := TRUE;
               RelWrite : Bool := FALSE;
            END_STRUCT;
            V_SerialNumber : Struct
               Text : String[64];
               Index : Int := 21;
               Subindex : Int := 0;
               Length : Int := 12;
               BlockStat : DWord;
               IOLStat : DWord;
               RelRead : Bool := TRUE;
               RelWrite : Bool := FALSE;
            END_STRUCT;
            V_HardwareRevision : Struct
               Text : String[64];
               Index : Int := 22;
               Subindex : Int := 0;
               Length : Int := 2;
               BlockStat : DWord;
               IOLStat : DWord;
               RelRead : Bool := TRUE;
               RelWrite : Bool := FALSE;
            END_STRUCT;
            V_FirmwareRevision : Struct
               Text : String[64];
               Index : Int := 23;
               Subindex : Int := 0;
               Length : Int := 5;
               BlockStat : DWord;
               IOLStat : DWord;
               RelRead : Bool := TRUE;
               RelWrite : Bool := FALSE;
            END_STRUCT;
         END_STRUCT;
         ApplicationSpecificTag : Struct
            V_ApplicationSpecificTag : Struct
               Text : String[64];
               Index : Int := 24;
               Subindex : Int := 0;
               Length : Int := 32;
               BlockStat : DWord;
               IOLStat : DWord;
               RelRead : Bool := TRUE;
               RelWrite : Bool := TRUE;
            END_STRUCT;
            V_FunctionTag : Struct
               Text : String[64];
               Index : Int := 25;
               Subindex : Int := 0;
               Length : Int := 0;
               BlockStat : DWord;
               IOLStat : DWord;
               RelRead : Bool := FALSE;
               RelWrite : Bool := FALSE;
            END_STRUCT;
            V_LocationTag : Struct
               Text : String[64];
               Index : Int := 26;
               Subindex : Int := 0;
               Length : Int := 0;
               BlockStat : DWord;
               IOLStat : DWord;
               RelRead : Bool := FALSE;
               RelWrite : Bool := FALSE;
            END_STRUCT;
         END_STRUCT;
         DeviceParameters : Struct
            Parameter_01 : Struct
               V_DeviceAccessLocks : Int := 0;
               Byte02 : Byte := BYTE#16#00;
               Byte03 : Byte := BYTE#16#00;
               Index : Int := 12;
               Subindex : Int := 0;
               Length : Int := 2;
               BlockStat : DWord;
               IOLStat : DWord;
               RelRead : Bool := TRUE;
               RelWrite : Bool := TRUE;
            END_STRUCT;
            Parameter_02 : Struct
               V_DeviceStatus : Byte := BYTE#16#00;
               Byte01 : Byte := BYTE#16#00;
               Byte02 : Byte := BYTE#16#00;
               Byte03 : Byte := BYTE#16#00;
               Index : Int := 36;
               Subindex : Int := 0;
               Length : Int := 1;
               BlockStat : DWord;
               IOLStat : DWord;
               RelRead : Bool := TRUE;
               RelWrite : Bool := FALSE;
            END_STRUCT;
            Parameter_03 : Struct
               V_BitCoded_ActiveEvents : DWord := DWORD#16#0000_0000;
               Index : Int := 545;
               Subindex : Int := 0;
               Length : Int := 4;
               BlockStat : DWord;
               IOLStat : DWord;
               RelRead : Bool := TRUE;
               RelWrite : Bool := FALSE;
            END_STRUCT;
            Parameter_04 : Struct
               V_ParaConfigFaultCollec : DInt := DINT#0;
               Index : Int := 546;
               Subindex : Int := 0;
               Length : Int := 4;
               BlockStat : DWord;
               IOLStat : DWord;
               RelRead : Bool := TRUE;
               RelWrite : Bool := FALSE;
            END_STRUCT;
            Parameter_05 : Struct
               V_EquipmentSpecificID : Byte := BYTE#16#00;
               Byte01 : Byte := BYTE#16#00;
               Byte02 : Byte := BYTE#16#00;
               Byte03 : Byte := BYTE#16#00;
               Index : Int := 688;
               Subindex : Int := 0;
               Length : Int := 1;
               BlockStat : DWord;
               IOLStat : DWord;
               RelRead : Bool := TRUE;
               RelWrite : Bool := TRUE;
            END_STRUCT;
            Parameter_06 : Struct
               V_X1_0_DO1Sub1 : Byte := BYTE#16#00;
               Byte01 : Byte := BYTE#16#00;
               Byte02 : Byte := BYTE#16#00;
               Byte03 : Byte := BYTE#16#00;
               Index : Int := 15000;
               Subindex : Int := 1;
               Length : Int := 1;
               BlockStat : DWord;
               IOLStat : DWord;
               RelRead : Bool := TRUE;
               RelWrite : Bool := TRUE;
            END_STRUCT;
            Parameter_07 : Struct
               V_X1_0_DO2Sub2 : Byte := BYTE#16#00;
               Byte01 : Byte := BYTE#16#00;
               Byte02 : Byte := BYTE#16#00;
               Byte03 : Byte := BYTE#16#00;
               Index : Int := 15000;
               Subindex : Int := 2;
               Length : Int := 1;
               BlockStat : DWord;
               IOLStat : DWord;
               RelRead : Bool := TRUE;
               RelWrite : Bool := TRUE;
            END_STRUCT;
            Parameter_08 : Struct
               V_X1_1_DO1Sub3 : Byte := BYTE#16#00;
               Byte01 : Byte := BYTE#16#00;
               Byte02 : Byte := BYTE#16#00;
               Byte03 : Byte := BYTE#16#00;
               Index : Int := 15000;
               Subindex : Int := 3;
               Length : Int := 1;
               BlockStat : DWord;
               IOLStat : DWord;
               RelRead : Bool := TRUE;
               RelWrite : Bool := TRUE;
            END_STRUCT;
            Parameter_09 : Struct
               V_X1_1_DO2Sub4 : Byte := BYTE#16#00;
               Byte01 : Byte := BYTE#16#00;
               Byte02 : Byte := BYTE#16#00;
               Byte03 : Byte := BYTE#16#00;
               Index : Int := 15000;
               Subindex : Int := 4;
               Length : Int := 1;
               BlockStat : DWord;
               IOLStat : DWord;
               RelRead : Bool := TRUE;
               RelWrite : Bool := TRUE;
            END_STRUCT;
            Parameter_10 : Struct
               V_X1_2_DO1Sub5 : Byte := BYTE#16#00;
               Byte01 : Byte := BYTE#16#00;
               Byte02 : Byte := BYTE#16#00;
               Byte03 : Byte := BYTE#16#00;
               Index : Int := 15000;
               Subindex : Int := 5;
               Length : Int := 1;
               BlockStat : DWord;
               IOLStat : DWord;
               RelRead : Bool := TRUE;
               RelWrite : Bool := TRUE;
            END_STRUCT;
            Parameter_11 : Struct
               V_X1_2_DO2Sub6 : Byte := BYTE#16#00;
               Byte01 : Byte := BYTE#16#00;
               Byte02 : Byte := BYTE#16#00;
               Byte03 : Byte := BYTE#16#00;
               Index : Int := 15000;
               Subindex : Int := 6;
               Length : Int := 1;
               BlockStat : DWord;
               IOLStat : DWord;
               RelRead : Bool := TRUE;
               RelWrite : Bool := TRUE;
            END_STRUCT;
            Parameter_12 : Struct
               V_X1_3_DO1Sub7 : Byte := BYTE#16#00;
               Byte01 : Byte := BYTE#16#00;
               Byte02 : Byte := BYTE#16#00;
               Byte03 : Byte := BYTE#16#00;
               Index : Int := 15000;
               Subindex : Int := 7;